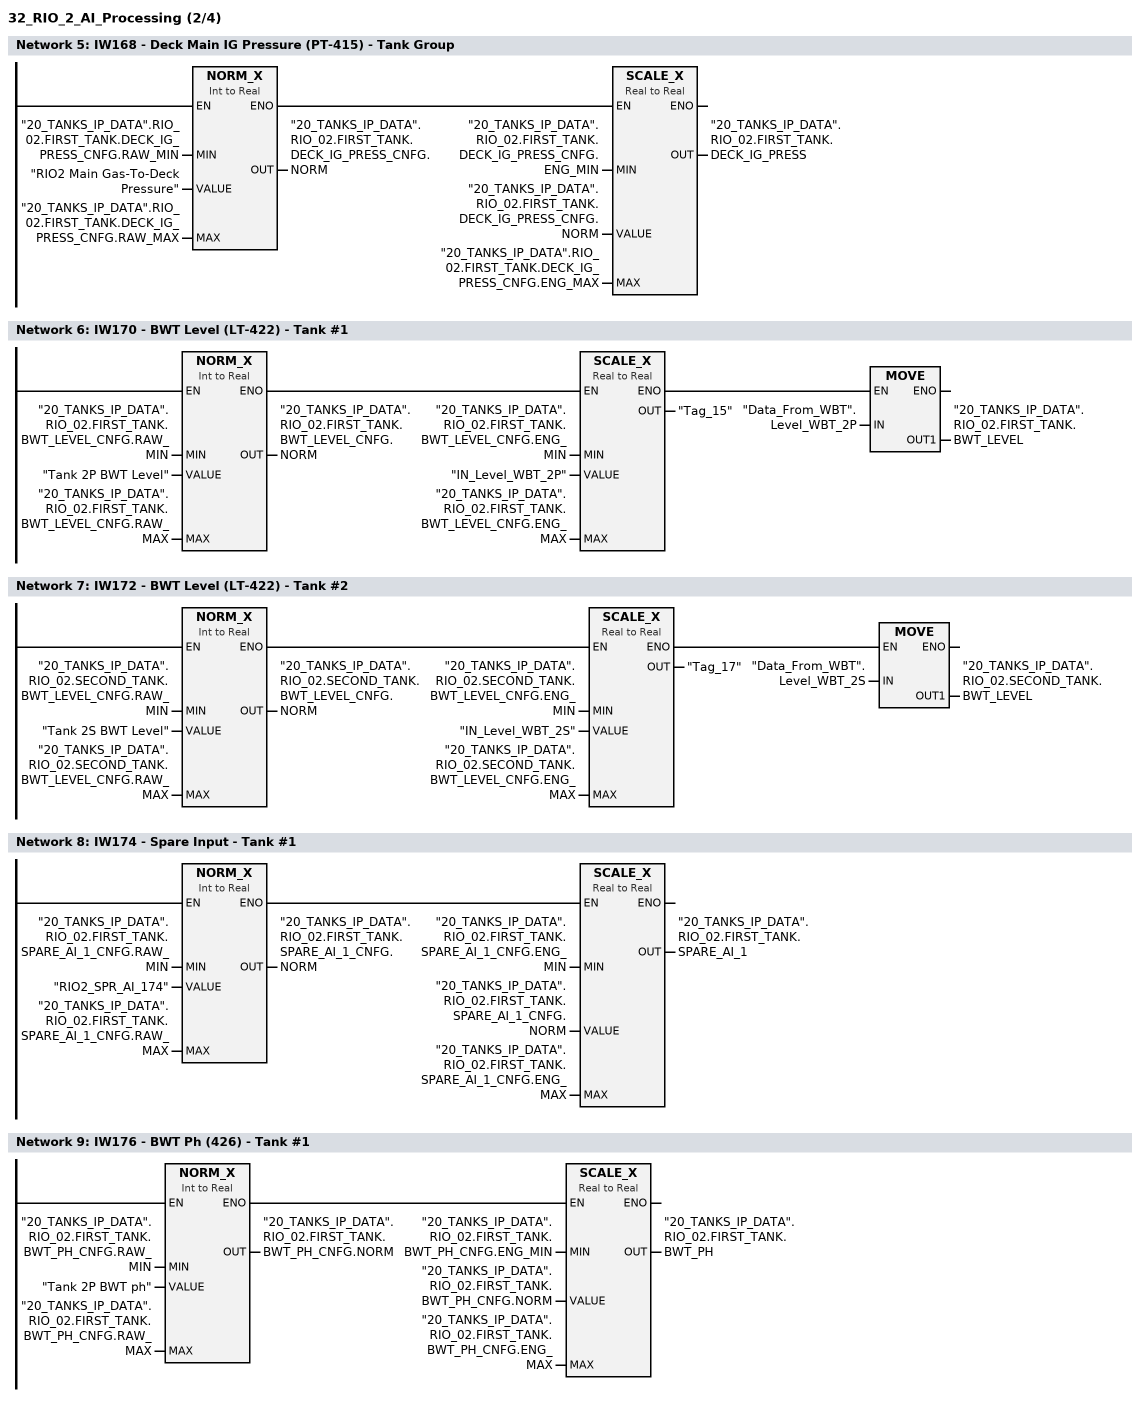
   RUNG wire#powerrail
      { S7_Templates := "[SrcType := Int, DestType := Real]" } Normalize(min := "20_TANKS_IP_DATA".RIO_02.FIRST_TANK.DECK_IG_PRESS_CNFG.RAW_MIN, value := "RIO2 Main Gas-To-Deck Pressure", max := "20_TANKS_IP_DATA".RIO_02.FIRST_TANK.DECK_IG_PRESS_CNFG.RAW_MAX, out => "20_TANKS_IP_DATA".RIO_02.FIRST_TANK.DECK_IG_PRESS_CNFG.NORM)
      { S7_Templates := "[SrcType := Real, DestType := Real]" } Scale(min := "20_TANKS_IP_DATA".RIO_02.FIRST_TANK.DECK_IG_PRESS_CNFG.ENG_MIN, value := "20_TANKS_IP_DATA".RIO_02.FIRST_TANK.DECK_IG_PRESS_CNFG.NORM, max := "20_TANKS_IP_DATA".RIO_02.FIRST_TANK.DECK_IG_PRESS_CNFG.ENG_MAX, out => "20_TANKS_IP_DATA".RIO_02.FIRST_TANK.DECK_IG_PRESS)
   END_RUNG
   // the same network as SCL:
   "20_TANKS_IP_DATA".RIO_02.FIRST_TANK.DECK_IG_PRESS_CNFG.NORM := NORM_X(MIN := "20_TANKS_IP_DATA".RIO_02.FIRST_TANK.DECK_IG_PRESS_CNFG.RAW_MIN, VALUE := "RIO2 Main Gas-To-Deck Pressure", MAX := "20_TANKS_IP_DATA".RIO_02.FIRST_TANK.DECK_IG_PRESS_CNFG.RAW_MAX);
   "20_TANKS_IP_DATA".RIO_02.FIRST_TANK.DECK_IG_PRESS := SCALE_X(MIN := "20_TANKS_IP_DATA".RIO_02.FIRST_TANK.DECK_IG_PRESS_CNFG.ENG_MIN, VALUE := "20_TANKS_IP_DATA".RIO_02.FIRST_TANK.DECK_IG_PRESS_CNFG.NORM, MAX := "20_TANKS_IP_DATA".RIO_02.FIRST_TANK.DECK_IG_PRESS_CNFG.ENG_MAX);
END_REGION

REGION Network 6: IW170 - BWT Level (LT-422) - Tank #1
   RUNG wire#powerrail
      { S7_Templates := "[SrcType := Int, DestType := Real]" } Normalize(min := "20_TANKS_IP_DATA".RIO_02.FIRST_TANK.BWT_LEVEL_CNFG.RAW_MIN, value := "Tank 2P BWT Level", max := "20_TANKS_IP_DATA".RIO_02.FIRST_TANK.BWT_LEVEL_CNFG.RAW_MAX, out => "20_TANKS_IP_DATA".RIO_02.FIRST_TANK.BWT_LEVEL_CNFG.NORM)
      { S7_Templates := "[SrcType := Real, DestType := Real]" } Scale(min := "20_TANKS_IP_DATA".RIO_02.FIRST_TANK.BWT_LEVEL_CNFG.ENG_MIN, value := "IN_Level_WBT_2P", max := "20_TANKS_IP_DATA".RIO_02.FIRST_TANK.BWT_LEVEL_CNFG.ENG_MAX, out => "Tag_15")
      Move(in := "Data_From_WBT".Level_WBT_2P, out1 => "20_TANKS_IP_DATA".RIO_02.FIRST_TANK.BWT_LEVEL)
   END_RUNG
   // the same network as SCL:
   "20_TANKS_IP_DATA".RIO_02.FIRST_TANK.BWT_LEVEL_CNFG.NORM := NORM_X(MIN := "20_TANKS_IP_DATA".RIO_02.FIRST_TANK.BWT_LEVEL_CNFG.RAW_MIN, VALUE := "Tank 2P BWT Level", MAX := "20_TANKS_IP_DATA".RIO_02.FIRST_TANK.BWT_LEVEL_CNFG.RAW_MAX);
   "Tag_15" := SCALE_X(MIN := "20_TANKS_IP_DATA".RIO_02.FIRST_TANK.BWT_LEVEL_CNFG.ENG_MIN, VALUE := "IN_Level_WBT_2P", MAX := "20_TANKS_IP_DATA".RIO_02.FIRST_TANK.BWT_LEVEL_CNFG.ENG_MAX);
   "20_TANKS_IP_DATA".RIO_02.FIRST_TANK.BWT_LEVEL := "Data_From_WBT".Level_WBT_2P;
END_REGION

REGION Network 7: IW172 - BWT Level (LT-422) - Tank #2
   RUNG wire#powerrail
      { S7_Templates := "[SrcType := Int, DestType := Real]" } Normalize(min := "20_TANKS_IP_DATA".RIO_02.SECOND_TANK.BWT_LEVEL_CNFG.RAW_MIN, value := "Tank 2S BWT Level", max := "20_TANKS_IP_DATA".RIO_02.SECOND_TANK.BWT_LEVEL_CNFG.RAW_MAX, out => "20_TANKS_IP_DATA".RIO_02.SECOND_TANK.BWT_LEVEL_CNFG.NORM)
      { S7_Templates := "[SrcType := Real, DestType := Real]" } Scale(min := "20_TANKS_IP_DATA".RIO_02.SECOND_TANK.BWT_LEVEL_CNFG.ENG_MIN, value := "IN_Level_WBT_2S", max := "20_TANKS_IP_DATA".RIO_02.SECOND_TANK.BWT_LEVEL_CNFG.ENG_MAX, out => "Tag_17")
      Move(in := "Data_From_WBT".Level_WBT_2S, out1 => "20_TANKS_IP_DATA".RIO_02.SECOND_TANK.BWT_LEVEL)
   END_RUNG
   // the same network as SCL:
   "20_TANKS_IP_DATA".RIO_02.SECOND_TANK.BWT_LEVEL_CNFG.NORM := NORM_X(MIN := "20_TANKS_IP_DATA".RIO_02.SECOND_TANK.BWT_LEVEL_CNFG.RAW_MIN, VALUE := "Tank 2S BWT Level", MAX := "20_TANKS_IP_DATA".RIO_02.SECOND_TANK.BWT_LEVEL_CNFG.RAW_MAX);
   "Tag_17" := SCALE_X(MIN := "20_TANKS_IP_DATA".RIO_02.SECOND_TANK.BWT_LEVEL_CNFG.ENG_MIN, VALUE := "IN_Level_WBT_2S", MAX := "20_TANKS_IP_DATA".RIO_02.SECOND_TANK.BWT_LEVEL_CNFG.ENG_MAX);
   "20_TANKS_IP_DATA".RIO_02.SECOND_TANK.BWT_LEVEL := "Data_From_WBT".Level_WBT_2S;
END_REGION

REGION Network 8: IW174 - Spare Input - Tank #1
   RUNG wire#powerrail
      { S7_Templates := "[SrcType := Int, DestType := Real]" } Normalize(min := "20_TANKS_IP_DATA".RIO_02.FIRST_TANK.SPARE_AI_1_CNFG.RAW_MIN, value := "RIO2_SPR_AI_174", max := "20_TANKS_IP_DATA".RIO_02.FIRST_TANK.SPARE_AI_1_CNFG.RAW_MAX, out => "20_TANKS_IP_DATA".RIO_02.FIRST_TANK.SPARE_AI_1_CNFG.NORM)
      { S7_Templates := "[SrcType := Real, DestType := Real]" } Scale(min := "20_TANKS_IP_DATA".RIO_02.FIRST_TANK.SPARE_AI_1_CNFG.ENG_MIN, value := "20_TANKS_IP_DATA".RIO_02.FIRST_TANK.SPARE_AI_1_CNFG.NORM, max := "20_TANKS_IP_DATA".RIO_02.FIRST_TANK.SPARE_AI_1_CNFG.ENG_MAX, out => "20_TANKS_IP_DATA".RIO_02.FIRST_TANK.SPARE_AI_1)
   END_RUNG
   // the same network as SCL:
   "20_TANKS_IP_DATA".RIO_02.FIRST_TANK.SPARE_AI_1_CNFG.NORM := NORM_X(MIN := "20_TANKS_IP_DATA".RIO_02.FIRST_TANK.SPARE_AI_1_CNFG.RAW_MIN, VALUE := "RIO2_SPR_AI_174", MAX := "20_TANKS_IP_DATA".RIO_02.FIRST_TANK.SPARE_AI_1_CNFG.RAW_MAX);
   "20_TANKS_IP_DATA".RIO_02.FIRST_TANK.SPARE_AI_1 := SCALE_X(MIN := "20_TANKS_IP_DATA".RIO_02.FIRST_TANK.SPARE_AI_1_CNFG.ENG_MIN, VALUE := "20_TANKS_IP_DATA".RIO_02.FIRST_TANK.SPARE_AI_1_CNFG.NORM, MAX := "20_TANKS_IP_DATA".RIO_02.FIRST_TANK.SPARE_AI_1_CNFG.ENG_MAX);
END_REGION

REGION Network 9: IW176 - BWT Ph (426) - Tank #1
   RUNG wire#powerrail
      { S7_Templates := "[SrcType := Int, DestType := Real]" } Normalize(min := "20_TANKS_IP_DATA".RIO_02.FIRST_TANK.BWT_PH_CNFG.RAW_MIN, value := "Tank 2P BWT ph", max := "20_TANKS_IP_DATA".RIO_02.FIRST_TANK.BWT_PH_CNFG.RAW_MAX, out => "20_TANKS_IP_DATA".RIO_02.FIRST_TANK.BWT_PH_CNFG.NORM)
      { S7_Templates := "[SrcType := Real, DestType := Real]" } Scale(min := "20_TANKS_IP_DATA".RIO_02.FIRST_TANK.BWT_PH_CNFG.ENG_MIN, value := "20_TANKS_IP_DATA".RIO_02.FIRST_TANK.BWT_PH_CNFG.NORM, max := "20_TANKS_IP_DATA".RIO_02.FIRST_TANK.BWT_PH_CNFG.ENG_MAX, out => "20_TANKS_IP_DATA".RIO_02.FIRST_TANK.BWT_PH)
   END_RUNG
   // the same network as SCL:
   "20_TANKS_IP_DATA".RIO_02.FIRST_TANK.BWT_PH_CNFG.NORM := NORM_X(MIN := "20_TANKS_IP_DATA".RIO_02.FIRST_TANK.BWT_PH_CNFG.RAW_MIN, VALUE := "Tank 2P BWT ph", MAX := "20_TANKS_IP_DATA".RIO_02.FIRST_TANK.BWT_PH_CNFG.RAW_MAX);
   "20_TANKS_IP_DATA".RIO_02.FIRST_TANK.BWT_PH := SCALE_X(MIN := "20_TANKS_IP_DATA".RIO_02.FIRST_TANK.BWT_PH_CNFG.ENG_MIN, VALUE := "20_TANKS_IP_DATA".RIO_02.FIRST_TANK.BWT_PH_CNFG.NORM, MAX := "20_TANKS_IP_DATA".RIO_02.FIRST_TANK.BWT_PH_CNFG.ENG_MAX);
END_REGION

REGION Network 10: IW178 - BWT Temperature (426) - Tank #1
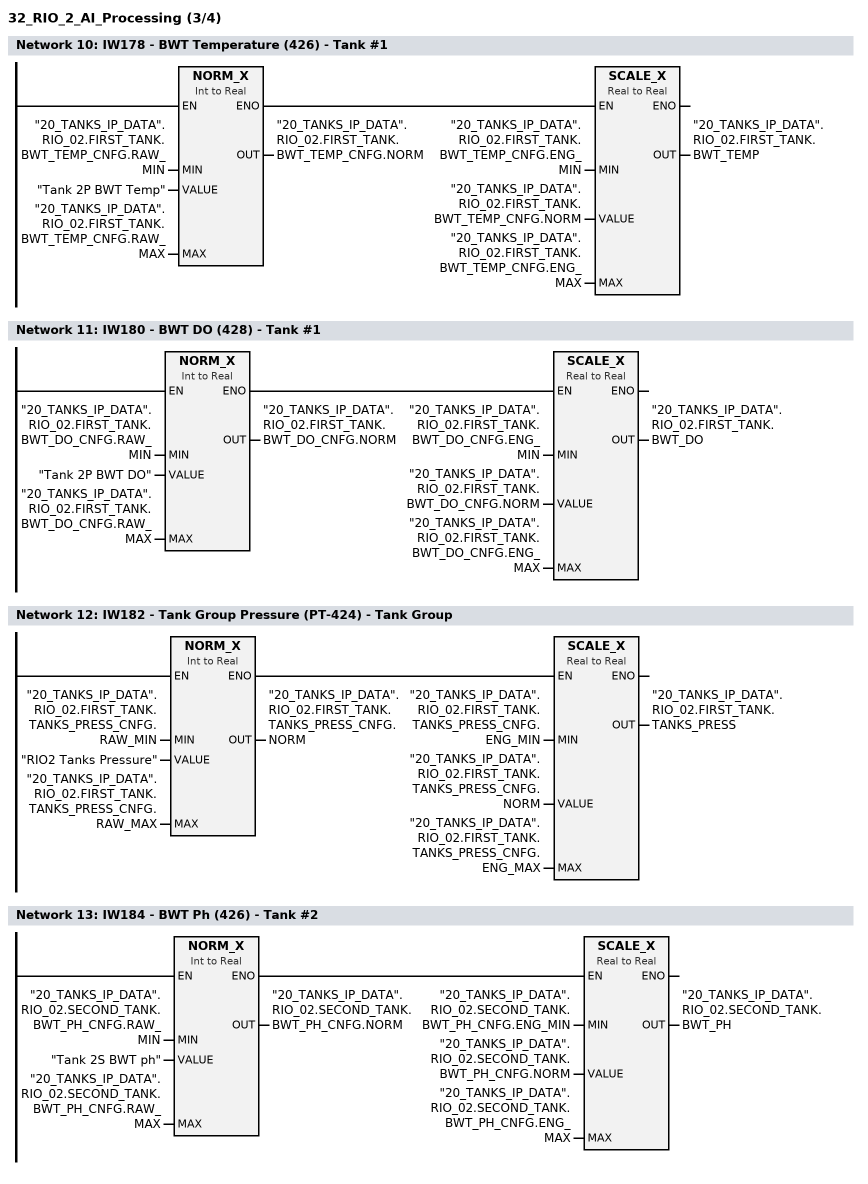
   RUNG wire#powerrail
      { S7_Templates := "[SrcType := Int, DestType := Real]" } Normalize(min := "20_TANKS_IP_DATA".RIO_02.FIRST_TANK.BWT_TEMP_CNFG.RAW_MIN, value := "Tank 2P BWT Temp", max := "20_TANKS_IP_DATA".RIO_02.FIRST_TANK.BWT_TEMP_CNFG.RAW_MAX, out => "20_TANKS_IP_DATA".RIO_02.FIRST_TANK.BWT_TEMP_CNFG.NORM)
      { S7_Templates := "[SrcType := Real, DestType := Real]" } Scale(min := "20_TANKS_IP_DATA".RIO_02.FIRST_TANK.BWT_TEMP_CNFG.ENG_MIN, value := "20_TANKS_IP_DATA".RIO_02.FIRST_TANK.BWT_TEMP_CNFG.NORM, max := "20_TANKS_IP_DATA".RIO_02.FIRST_TANK.BWT_TEMP_CNFG.ENG_MAX, out => "20_TANKS_IP_DATA".RIO_02.FIRST_TANK.BWT_TEMP)
   END_RUNG
   // the same network as SCL:
   "20_TANKS_IP_DATA".RIO_02.FIRST_TANK.BWT_TEMP_CNFG.NORM := NORM_X(MIN := "20_TANKS_IP_DATA".RIO_02.FIRST_TANK.BWT_TEMP_CNFG.RAW_MIN, VALUE := "Tank 2P BWT Temp", MAX := "20_TANKS_IP_DATA".RIO_02.FIRST_TANK.BWT_TEMP_CNFG.RAW_MAX);
   "20_TANKS_IP_DATA".RIO_02.FIRST_TANK.BWT_TEMP := SCALE_X(MIN := "20_TANKS_IP_DATA".RIO_02.FIRST_TANK.BWT_TEMP_CNFG.ENG_MIN, VALUE := "20_TANKS_IP_DATA".RIO_02.FIRST_TANK.BWT_TEMP_CNFG.NORM, MAX := "20_TANKS_IP_DATA".RIO_02.FIRST_TANK.BWT_TEMP_CNFG.ENG_MAX);
END_REGION

REGION Network 11: IW180 - BWT DO (428) - Tank #1
   RUNG wire#powerrail
      { S7_Templates := "[SrcType := Int, DestType := Real]" } Normalize(min := "20_TANKS_IP_DATA".RIO_02.FIRST_TANK.BWT_DO_CNFG.RAW_MIN, value := "Tank 2P BWT DO", max := "20_TANKS_IP_DATA".RIO_02.FIRST_TANK.BWT_DO_CNFG.RAW_MAX, out => "20_TANKS_IP_DATA".RIO_02.FIRST_TANK.BWT_DO_CNFG.NORM)
      { S7_Templates := "[SrcType := Real, DestType := Real]" } Scale(min := "20_TANKS_IP_DATA".RIO_02.FIRST_TANK.BWT_DO_CNFG.ENG_MIN, value := "20_TANKS_IP_DATA".RIO_02.FIRST_TANK.BWT_DO_CNFG.NORM, max := "20_TANKS_IP_DATA".RIO_02.FIRST_TANK.BWT_DO_CNFG.ENG_MAX, out => "20_TANKS_IP_DATA".RIO_02.FIRST_TANK.BWT_DO)
   END_RUNG
   // the same network as SCL:
   "20_TANKS_IP_DATA".RIO_02.FIRST_TANK.BWT_DO_CNFG.NORM := NORM_X(MIN := "20_TANKS_IP_DATA".RIO_02.FIRST_TANK.BWT_DO_CNFG.RAW_MIN, VALUE := "Tank 2P BWT DO", MAX := "20_TANKS_IP_DATA".RIO_02.FIRST_TANK.BWT_DO_CNFG.RAW_MAX);
   "20_TANKS_IP_DATA".RIO_02.FIRST_TANK.BWT_DO := SCALE_X(MIN := "20_TANKS_IP_DATA".RIO_02.FIRST_TANK.BWT_DO_CNFG.ENG_MIN, VALUE := "20_TANKS_IP_DATA".RIO_02.FIRST_TANK.BWT_DO_CNFG.NORM, MAX := "20_TANKS_IP_DATA".RIO_02.FIRST_TANK.BWT_DO_CNFG.ENG_MAX);
END_REGION

REGION Network 12: IW182 - Tank Group Pressure (PT-424) - Tank Group
   RUNG wire#powerrail
      { S7_Templates := "[SrcType := Int, DestType := Real]" } Normalize(min := "20_TANKS_IP_DATA".RIO_02.FIRST_TANK.TANKS_PRESS_CNFG.RAW_MIN, value := "RIO2 Tanks Pressure", max := "20_TANKS_IP_DATA".RIO_02.FIRST_TANK.TANKS_PRESS_CNFG.RAW_MAX, out => "20_TANKS_IP_DATA".RIO_02.FIRST_TANK.TANKS_PRESS_CNFG.NORM)
      { S7_Templates := "[SrcType := Real, DestType := Real]" } Scale(min := "20_TANKS_IP_DATA".RIO_02.FIRST_TANK.TANKS_PRESS_CNFG.ENG_MIN, value := "20_TANKS_IP_DATA".RIO_02.FIRST_TANK.TANKS_PRESS_CNFG.NORM, max := "20_TANKS_IP_DATA".RIO_02.FIRST_TANK.TANKS_PRESS_CNFG.ENG_MAX, out => "20_TANKS_IP_DATA".RIO_02.FIRST_TANK.TANKS_PRESS)
   END_RUNG
   // the same network as SCL:
   "20_TANKS_IP_DATA".RIO_02.FIRST_TANK.TANKS_PRESS_CNFG.NORM := NORM_X(MIN := "20_TANKS_IP_DATA".RIO_02.FIRST_TANK.TANKS_PRESS_CNFG.RAW_MIN, VALUE := "RIO2 Tanks Pressure", MAX := "20_TANKS_IP_DATA".RIO_02.FIRST_TANK.TANKS_PRESS_CNFG.RAW_MAX);
   "20_TANKS_IP_DATA".RIO_02.FIRST_TANK.TANKS_PRESS := SCALE_X(MIN := "20_TANKS_IP_DATA".RIO_02.FIRST_TANK.TANKS_PRESS_CNFG.ENG_MIN, VALUE := "20_TANKS_IP_DATA".RIO_02.FIRST_TANK.TANKS_PRESS_CNFG.NORM, MAX := "20_TANKS_IP_DATA".RIO_02.FIRST_TANK.TANKS_PRESS_CNFG.ENG_MAX);
END_REGION

REGION Network 13: IW184 - BWT Ph (426) - Tank #2
   RUNG wire#powerrail
      { S7_Templates := "[SrcType := Int, DestType := Real]" } Normalize(min := "20_TANKS_IP_DATA".RIO_02.SECOND_TANK.BWT_PH_CNFG.RAW_MIN, value := "Tank 2S BWT ph", max := "20_TANKS_IP_DATA".RIO_02.SECOND_TANK.BWT_PH_CNFG.RAW_MAX, out => "20_TANKS_IP_DATA".RIO_02.SECOND_TANK.BWT_PH_CNFG.NORM)
      { S7_Templates := "[SrcType := Real, DestType := Real]" } Scale(min := "20_TANKS_IP_DATA".RIO_02.SECOND_TANK.BWT_PH_CNFG.ENG_MIN, value := "20_TANKS_IP_DATA".RIO_02.SECOND_TANK.BWT_PH_CNFG.NORM, max := "20_TANKS_IP_DATA".RIO_02.SECOND_TANK.BWT_PH_CNFG.ENG_MAX, out => "20_TANKS_IP_DATA".RIO_02.SECOND_TANK.BWT_PH)
   END_RUNG
   // the same network as SCL:
   "20_TANKS_IP_DATA".RIO_02.SECOND_TANK.BWT_PH_CNFG.NORM := NORM_X(MIN := "20_TANKS_IP_DATA".RIO_02.SECOND_TANK.BWT_PH_CNFG.RAW_MIN, VALUE := "Tank 2S BWT ph", MAX := "20_TANKS_IP_DATA".RIO_02.SECOND_TANK.BWT_PH_CNFG.RAW_MAX);
   "20_TANKS_IP_DATA".RIO_02.SECOND_TANK.BWT_PH := SCALE_X(MIN := "20_TANKS_IP_DATA".RIO_02.SECOND_TANK.BWT_PH_CNFG.ENG_MIN, VALUE := "20_TANKS_IP_DATA".RIO_02.SECOND_TANK.BWT_PH_CNFG.NORM, MAX := "20_TANKS_IP_DATA".RIO_02.SECOND_TANK.BWT_PH_CNFG.ENG_MAX);
END_REGION

REGION Network 14: IW186 - BWT Temperature (426) - Tank #2
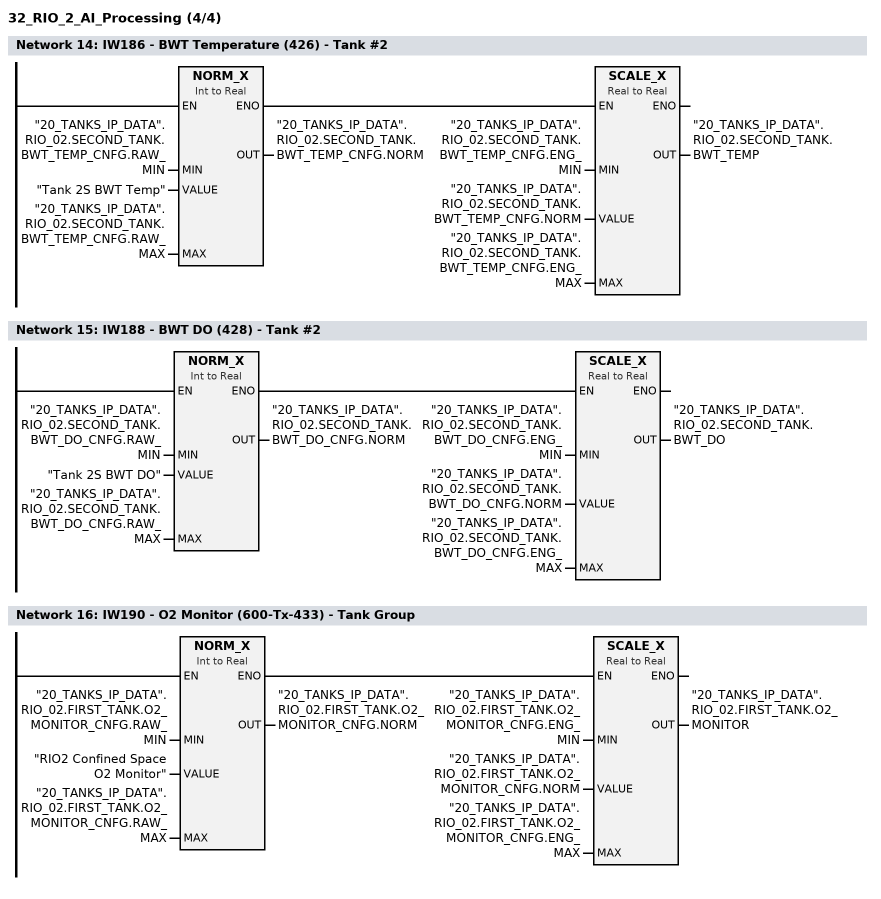
   RUNG wire#powerrail
      { S7_Templates := "[SrcType := Int, DestType := Real]" } Normalize(min := "20_TANKS_IP_DATA".RIO_02.SECOND_TANK.BWT_TEMP_CNFG.RAW_MIN, value := "Tank 2S BWT Temp", max := "20_TANKS_IP_DATA".RIO_02.SECOND_TANK.BWT_TEMP_CNFG.RAW_MAX, out => "20_TANKS_IP_DATA".RIO_02.SECOND_TANK.BWT_TEMP_CNFG.NORM)
      { S7_Templates := "[SrcType := Real, DestType := Real]" } Scale(min := "20_TANKS_IP_DATA".RIO_02.SECOND_TANK.BWT_TEMP_CNFG.ENG_MIN, value := "20_TANKS_IP_DATA".RIO_02.SECOND_TANK.BWT_TEMP_CNFG.NORM, max := "20_TANKS_IP_DATA".RIO_02.SECOND_TANK.BWT_TEMP_CNFG.ENG_MAX, out => "20_TANKS_IP_DATA".RIO_02.SECOND_TANK.BWT_TEMP)
   END_RUNG
   // the same network as SCL:
   "20_TANKS_IP_DATA".RIO_02.SECOND_TANK.BWT_TEMP_CNFG.NORM := NORM_X(MIN := "20_TANKS_IP_DATA".RIO_02.SECOND_TANK.BWT_TEMP_CNFG.RAW_MIN, VALUE := "Tank 2S BWT Temp", MAX := "20_TANKS_IP_DATA".RIO_02.SECOND_TANK.BWT_TEMP_CNFG.RAW_MAX);
   "20_TANKS_IP_DATA".RIO_02.SECOND_TANK.BWT_TEMP := SCALE_X(MIN := "20_TANKS_IP_DATA".RIO_02.SECOND_TANK.BWT_TEMP_CNFG.ENG_MIN, VALUE := "20_TANKS_IP_DATA".RIO_02.SECOND_TANK.BWT_TEMP_CNFG.NORM, MAX := "20_TANKS_IP_DATA".RIO_02.SECOND_TANK.BWT_TEMP_CNFG.ENG_MAX);
END_REGION

REGION Network 15: IW188 - BWT DO (428) - Tank #2
   RUNG wire#powerrail
      { S7_Templates := "[SrcType := Int, DestType := Real]" } Normalize(min := "20_TANKS_IP_DATA".RIO_02.SECOND_TANK.BWT_DO_CNFG.RAW_MIN, value := "Tank 2S BWT DO", max := "20_TANKS_IP_DATA".RIO_02.SECOND_TANK.BWT_DO_CNFG.RAW_MAX, out => "20_TANKS_IP_DATA".RIO_02.SECOND_TANK.BWT_DO_CNFG.NORM)
      { S7_Templates := "[SrcType := Real, DestType := Real]" } Scale(min := "20_TANKS_IP_DATA".RIO_02.SECOND_TANK.BWT_DO_CNFG.ENG_MIN, value := "20_TANKS_IP_DATA".RIO_02.SECOND_TANK.BWT_DO_CNFG.NORM, max := "20_TANKS_IP_DATA".RIO_02.SECOND_TANK.BWT_DO_CNFG.ENG_MAX, out => "20_TANKS_IP_DATA".RIO_02.SECOND_TANK.BWT_DO)
   END_RUNG
   // the same network as SCL:
   "20_TANKS_IP_DATA".RIO_02.SECOND_TANK.BWT_DO_CNFG.NORM := NORM_X(MIN := "20_TANKS_IP_DATA".RIO_02.SECOND_TANK.BWT_DO_CNFG.RAW_MIN, VALUE := "Tank 2S BWT DO", MAX := "20_TANKS_IP_DATA".RIO_02.SECOND_TANK.BWT_DO_CNFG.RAW_MAX);
   "20_TANKS_IP_DATA".RIO_02.SECOND_TANK.BWT_DO := SCALE_X(MIN := "20_TANKS_IP_DATA".RIO_02.SECOND_TANK.BWT_DO_CNFG.ENG_MIN, VALUE := "20_TANKS_IP_DATA".RIO_02.SECOND_TANK.BWT_DO_CNFG.NORM, MAX := "20_TANKS_IP_DATA".RIO_02.SECOND_TANK.BWT_DO_CNFG.ENG_MAX);
END_REGION

REGION Network 16: IW190 - O2 Monitor (600-Tx-433) - Tank Group
   RUNG wire#powerrail
      { S7_Templates := "[SrcType := Int, DestType := Real]" } Normalize(min := "20_TANKS_IP_DATA".RIO_02.FIRST_TANK.O2_MONITOR_CNFG.RAW_MIN, value := "RIO2 Confined Space O2 Monitor", max := "20_TANKS_IP_DATA".RIO_02.FIRST_TANK.O2_MONITOR_CNFG.RAW_MAX, out => "20_TANKS_IP_DATA".RIO_02.FIRST_TANK.O2_MONITOR_CNFG.NORM)
      { S7_Templates := "[SrcType := Real, DestType := Real]" } Scale(min := "20_TANKS_IP_DATA".RIO_02.FIRST_TANK.O2_MONITOR_CNFG.ENG_MIN, value := "20_TANKS_IP_DATA".RIO_02.FIRST_TANK.O2_MONITOR_CNFG.NORM, max := "20_TANKS_IP_DATA".RIO_02.FIRST_TANK.O2_MONITOR_CNFG.ENG_MAX, out => "20_TANKS_IP_DATA".RIO_02.FIRST_TANK.O2_MONITOR)
   END_RUNG
   // the same network as SCL:
   "20_TANKS_IP_DATA".RIO_02.FIRST_TANK.O2_MONITOR_CNFG.NORM := NORM_X(MIN := "20_TANKS_IP_DATA".RIO_02.FIRST_TANK.O2_MONITOR_CNFG.RAW_MIN, VALUE := "RIO2 Confined Space O2 Monitor", MAX := "20_TANKS_IP_DATA".RIO_02.FIRST_TANK.O2_MONITOR_CNFG.RAW_MAX);
   "20_TANKS_IP_DATA".RIO_02.FIRST_TANK.O2_MONITOR := SCALE_X(MIN := "20_TANKS_IP_DATA".RIO_02.FIRST_TANK.O2_MONITOR_CNFG.ENG_MIN, VALUE := "20_TANKS_IP_DATA".RIO_02.FIRST_TANK.O2_MONITOR_CNFG.NORM, MAX := "20_TANKS_IP_DATA".RIO_02.FIRST_TANK.O2_MONITOR_CNFG.ENG_MAX);
END_REGION
END_FUNCTION

FUNCTION "33_RIO_3_AI_Processing" : Void   // FC33, LAD
TITLE = Analogue Input Processing (Tank 1 = 3P, Tank 2 = 3S)
{ S7_Optimized_Access := 'TRUE' }
AUTHOR : JRS
VERSION : 0.1
// To process raw inputs prior to code use
BEGIN

REGION Network 1: IW200 - USD Flow (FIT-418) - Tank #1
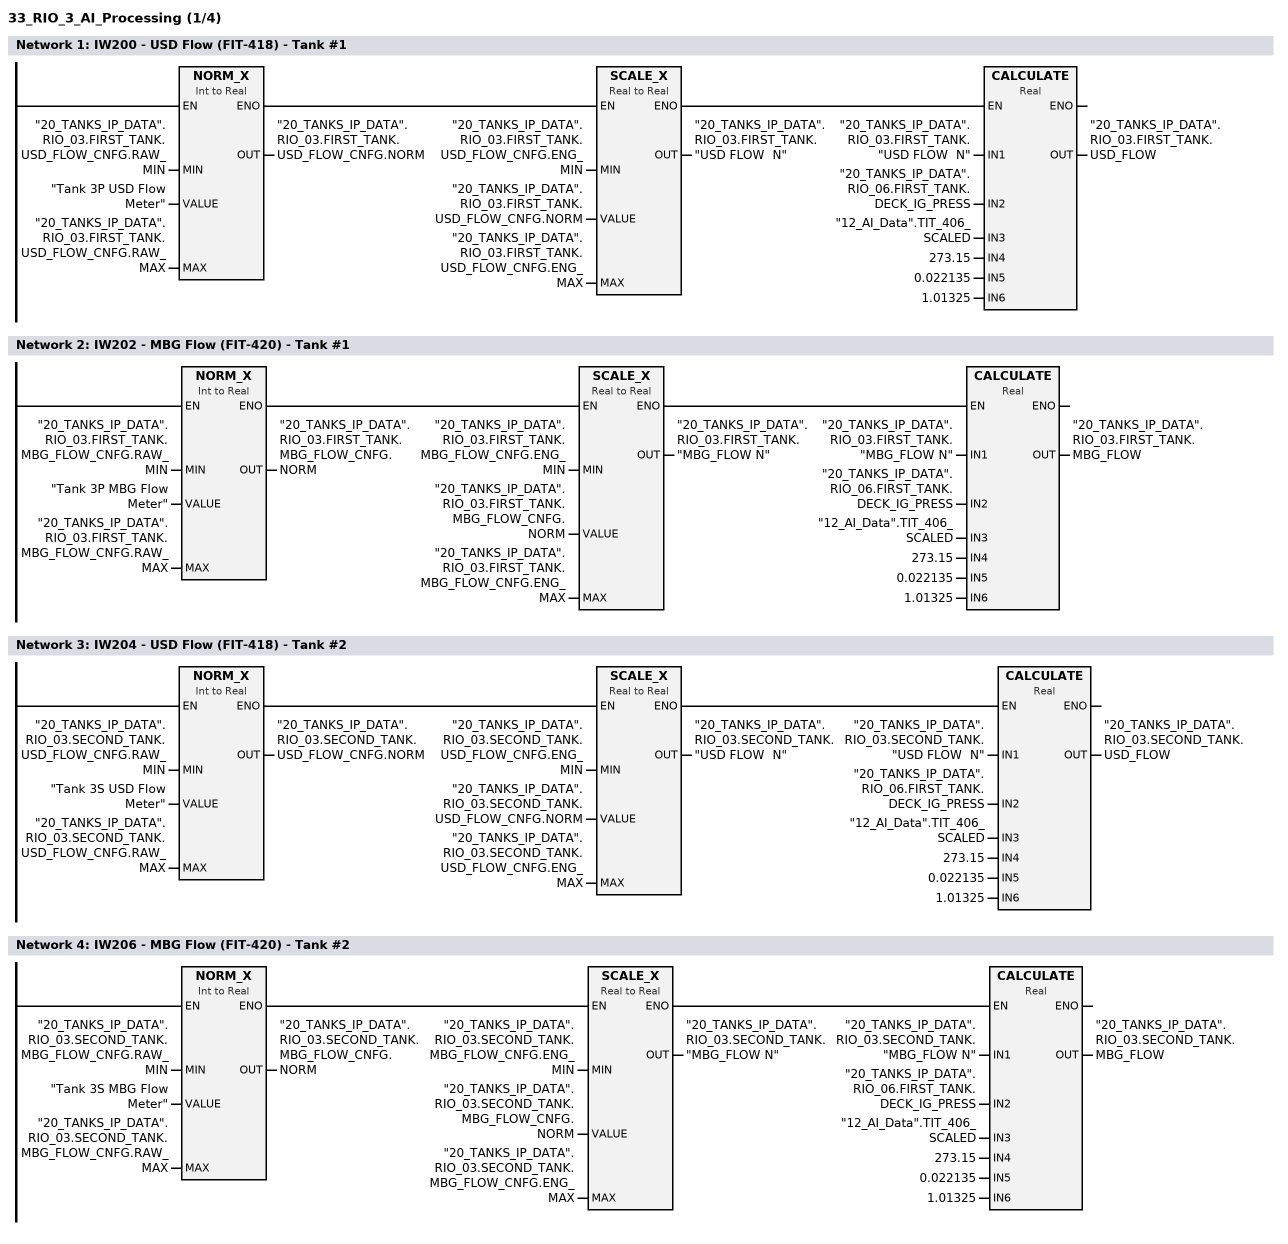
   RUNG wire#powerrail
      { S7_Templates := "[SrcType := Int, DestType := Real]" } Normalize(min := "20_TANKS_IP_DATA".RIO_03.FIRST_TANK.USD_FLOW_CNFG.RAW_MIN, value := "Tank 3P USD Flow Meter", max := "20_TANKS_IP_DATA".RIO_03.FIRST_TANK.USD_FLOW_CNFG.RAW_MAX, out => "20_TANKS_IP_DATA".RIO_03.FIRST_TANK.USD_FLOW_CNFG.NORM)
      { S7_Templates := "[SrcType := Real, DestType := Real]" } Scale(min := "20_TANKS_IP_DATA".RIO_03.FIRST_TANK.USD_FLOW_CNFG.ENG_MIN, value := "20_TANKS_IP_DATA".RIO_03.FIRST_TANK.USD_FLOW_CNFG.NORM, max := "20_TANKS_IP_DATA".RIO_03.FIRST_TANK.USD_FLOW_CNFG.ENG_MAX, out => "20_TANKS_IP_DATA".RIO_03.FIRST_TANK."USD FLOW  N")
      { S7_Templates := "SrcType := Real"; S7_Expression := "IN1*(IN2+IN6)/IN6*IN4/(IN3+IN4)" } Calculate(in1 := "20_TANKS_IP_DATA".RIO_03.FIRST_TANK."USD FLOW  N", in2 := "20_TANKS_IP_DATA".RIO_06.FIRST_TANK.DECK_IG_PRESS, in3 := "12_AI_Data".TIT_406_SCALED, in4 := 273.15, in5 := 0.022135, in6 := 1.01325, out => "20_TANKS_IP_DATA".RIO_03.FIRST_TANK.USD_FLOW)
   END_RUNG
   // the same network as SCL:
   "20_TANKS_IP_DATA".RIO_03.FIRST_TANK.USD_FLOW_CNFG.NORM := NORM_X(MIN := "20_TANKS_IP_DATA".RIO_03.FIRST_TANK.USD_FLOW_CNFG.RAW_MIN, VALUE := "Tank 3P USD Flow Meter", MAX := "20_TANKS_IP_DATA".RIO_03.FIRST_TANK.USD_FLOW_CNFG.RAW_MAX);
   "20_TANKS_IP_DATA".RIO_03.FIRST_TANK."USD FLOW  N" := SCALE_X(MIN := "20_TANKS_IP_DATA".RIO_03.FIRST_TANK.USD_FLOW_CNFG.ENG_MIN, VALUE := "20_TANKS_IP_DATA".RIO_03.FIRST_TANK.USD_FLOW_CNFG.NORM, MAX := "20_TANKS_IP_DATA".RIO_03.FIRST_TANK.USD_FLOW_CNFG.ENG_MAX);
   "20_TANKS_IP_DATA".RIO_03.FIRST_TANK.USD_FLOW := "20_TANKS_IP_DATA".RIO_03.FIRST_TANK."USD FLOW  N"*("20_TANKS_IP_DATA".RIO_06.FIRST_TANK.DECK_IG_PRESS+1.01325)/1.01325*273.15/("12_AI_Data".TIT_406_SCALED+273.15);
END_REGION

REGION Network 2: IW202 - MBG Flow (FIT-420) - Tank #1
   RUNG wire#powerrail
      { S7_Templates := "[SrcType := Int, DestType := Real]" } Normalize(min := "20_TANKS_IP_DATA".RIO_03.FIRST_TANK.MBG_FLOW_CNFG.RAW_MIN, value := "Tank 3P MBG Flow Meter", max := "20_TANKS_IP_DATA".RIO_03.FIRST_TANK.MBG_FLOW_CNFG.RAW_MAX, out => "20_TANKS_IP_DATA".RIO_03.FIRST_TANK.MBG_FLOW_CNFG.NORM)
      { S7_Templates := "[SrcType := Real, DestType := Real]" } Scale(min := "20_TANKS_IP_DATA".RIO_03.FIRST_TANK.MBG_FLOW_CNFG.ENG_MIN, value := "20_TANKS_IP_DATA".RIO_03.FIRST_TANK.MBG_FLOW_CNFG.NORM, max := "20_TANKS_IP_DATA".RIO_03.FIRST_TANK.MBG_FLOW_CNFG.ENG_MAX, out => "20_TANKS_IP_DATA".RIO_03.FIRST_TANK."MBG_FLOW N")
      { S7_Templates := "SrcType := Real"; S7_Expression := "IN1*(IN2+IN6)/IN6*IN4/(IN3+IN4)" } Calculate(in1 := "20_TANKS_IP_DATA".RIO_03.FIRST_TANK."MBG_FLOW N", in2 := "20_TANKS_IP_DATA".RIO_06.FIRST_TANK.DECK_IG_PRESS, in3 := "12_AI_Data".TIT_406_SCALED, in4 := 273.15, in5 := 0.022135, in6 := 1.01325, out => "20_TANKS_IP_DATA".RIO_03.FIRST_TANK.MBG_FLOW)
   END_RUNG
   // the same network as SCL:
   "20_TANKS_IP_DATA".RIO_03.FIRST_TANK.MBG_FLOW_CNFG.NORM := NORM_X(MIN := "20_TANKS_IP_DATA".RIO_03.FIRST_TANK.MBG_FLOW_CNFG.RAW_MIN, VALUE := "Tank 3P MBG Flow Meter", MAX := "20_TANKS_IP_DATA".RIO_03.FIRST_TANK.MBG_FLOW_CNFG.RAW_MAX);
   "20_TANKS_IP_DATA".RIO_03.FIRST_TANK."MBG_FLOW N" := SCALE_X(MIN := "20_TANKS_IP_DATA".RIO_03.FIRST_TANK.MBG_FLOW_CNFG.ENG_MIN, VALUE := "20_TANKS_IP_DATA".RIO_03.FIRST_TANK.MBG_FLOW_CNFG.NORM, MAX := "20_TANKS_IP_DATA".RIO_03.FIRST_TANK.MBG_FLOW_CNFG.ENG_MAX);
   "20_TANKS_IP_DATA".RIO_03.FIRST_TANK.MBG_FLOW := "20_TANKS_IP_DATA".RIO_03.FIRST_TANK."MBG_FLOW N"*("20_TANKS_IP_DATA".RIO_06.FIRST_TANK.DECK_IG_PRESS+1.01325)/1.01325*273.15/("12_AI_Data".TIT_406_SCALED+273.15);
END_REGION

REGION Network 3: IW204 - USD Flow (FIT-418) - Tank #2
   RUNG wire#powerrail
      { S7_Templates := "[SrcType := Int, DestType := Real]" } Normalize(min := "20_TANKS_IP_DATA".RIO_03.SECOND_TANK.USD_FLOW_CNFG.RAW_MIN, value := "Tank 3S USD Flow Meter", max := "20_TANKS_IP_DATA".RIO_03.SECOND_TANK.USD_FLOW_CNFG.RAW_MAX, out => "20_TANKS_IP_DATA".RIO_03.SECOND_TANK.USD_FLOW_CNFG.NORM)
      { S7_Templates := "[SrcType := Real, DestType := Real]" } Scale(min := "20_TANKS_IP_DATA".RIO_03.SECOND_TANK.USD_FLOW_CNFG.ENG_MIN, value := "20_TANKS_IP_DATA".RIO_03.SECOND_TANK.USD_FLOW_CNFG.NORM, max := "20_TANKS_IP_DATA".RIO_03.SECOND_TANK.USD_FLOW_CNFG.ENG_MAX, out => "20_TANKS_IP_DATA".RIO_03.SECOND_TANK."USD FLOW  N")
      { S7_Templates := "SrcType := Real"; S7_Expression := "IN1*(IN2+IN6)/IN6*IN4/(IN3+IN4)" } Calculate(in1 := "20_TANKS_IP_DATA".RIO_03.SECOND_TANK."USD FLOW  N", in2 := "20_TANKS_IP_DATA".RIO_06.FIRST_TANK.DECK_IG_PRESS, in3 := "12_AI_Data".TIT_406_SCALED, in4 := 273.15, in5 := 0.022135, in6 := 1.01325, out => "20_TANKS_IP_DATA".RIO_03.SECOND_TANK.USD_FLOW)
   END_RUNG
   // the same network as SCL:
   "20_TANKS_IP_DATA".RIO_03.SECOND_TANK.USD_FLOW_CNFG.NORM := NORM_X(MIN := "20_TANKS_IP_DATA".RIO_03.SECOND_TANK.USD_FLOW_CNFG.RAW_MIN, VALUE := "Tank 3S USD Flow Meter", MAX := "20_TANKS_IP_DATA".RIO_03.SECOND_TANK.USD_FLOW_CNFG.RAW_MAX);
   "20_TANKS_IP_DATA".RIO_03.SECOND_TANK."USD FLOW  N" := SCALE_X(MIN := "20_TANKS_IP_DATA".RIO_03.SECOND_TANK.USD_FLOW_CNFG.ENG_MIN, VALUE := "20_TANKS_IP_DATA".RIO_03.SECOND_TANK.USD_FLOW_CNFG.NORM, MAX := "20_TANKS_IP_DATA".RIO_03.SECOND_TANK.USD_FLOW_CNFG.ENG_MAX);
   "20_TANKS_IP_DATA".RIO_03.SECOND_TANK.USD_FLOW := "20_TANKS_IP_DATA".RIO_03.SECOND_TANK."USD FLOW  N"*("20_TANKS_IP_DATA".RIO_06.FIRST_TANK.DECK_IG_PRESS+1.01325)/1.01325*273.15/("12_AI_Data".TIT_406_SCALED+273.15);
END_REGION

REGION Network 4: IW206 - MBG Flow (FIT-420) - Tank #2
   RUNG wire#powerrail
      { S7_Templates := "[SrcType := Int, DestType := Real]" } Normalize(min := "20_TANKS_IP_DATA".RIO_03.SECOND_TANK.MBG_FLOW_CNFG.RAW_MIN, value := "Tank 3S MBG Flow Meter", max := "20_TANKS_IP_DATA".RIO_03.SECOND_TANK.MBG_FLOW_CNFG.RAW_MAX, out => "20_TANKS_IP_DATA".RIO_03.SECOND_TANK.MBG_FLOW_CNFG.NORM)
      { S7_Templates := "[SrcType := Real, DestType := Real]" } Scale(min := "20_TANKS_IP_DATA".RIO_03.SECOND_TANK.MBG_FLOW_CNFG.ENG_MIN, value := "20_TANKS_IP_DATA".RIO_03.SECOND_TANK.MBG_FLOW_CNFG.NORM, max := "20_TANKS_IP_DATA".RIO_03.SECOND_TANK.MBG_FLOW_CNFG.ENG_MAX, out => "20_TANKS_IP_DATA".RIO_03.SECOND_TANK."MBG_FLOW N")
      { S7_Templates := "SrcType := Real"; S7_Expression := "IN1*(IN2+IN6)/IN6*IN4/(IN3+IN4)" } Calculate(in1 := "20_TANKS_IP_DATA".RIO_03.SECOND_TANK."MBG_FLOW N", in2 := "20_TANKS_IP_DATA".RIO_06.FIRST_TANK.DECK_IG_PRESS, in3 := "12_AI_Data".TIT_406_SCALED, in4 := 273.15, in5 := 0.022135, in6 := 1.01325, out => "20_TANKS_IP_DATA".RIO_03.SECOND_TANK.MBG_FLOW)
   END_RUNG
   // the same network as SCL:
   "20_TANKS_IP_DATA".RIO_03.SECOND_TANK.MBG_FLOW_CNFG.NORM := NORM_X(MIN := "20_TANKS_IP_DATA".RIO_03.SECOND_TANK.MBG_FLOW_CNFG.RAW_MIN, VALUE := "Tank 3S MBG Flow Meter", MAX := "20_TANKS_IP_DATA".RIO_03.SECOND_TANK.MBG_FLOW_CNFG.RAW_MAX);
   "20_TANKS_IP_DATA".RIO_03.SECOND_TANK."MBG_FLOW N" := SCALE_X(MIN := "20_TANKS_IP_DATA".RIO_03.SECOND_TANK.MBG_FLOW_CNFG.ENG_MIN, VALUE := "20_TANKS_IP_DATA".RIO_03.SECOND_TANK.MBG_FLOW_CNFG.NORM, MAX := "20_TANKS_IP_DATA".RIO_03.SECOND_TANK.MBG_FLOW_CNFG.ENG_MAX);
   "20_TANKS_IP_DATA".RIO_03.SECOND_TANK.MBG_FLOW := "20_TANKS_IP_DATA".RIO_03.SECOND_TANK."MBG_FLOW N"*("20_TANKS_IP_DATA".RIO_06.FIRST_TANK.DECK_IG_PRESS+1.01325)/1.01325*273.15/("12_AI_Data".TIT_406_SCALED+273.15);
END_REGION

REGION Network 5: IW208 - Deck Main IG Pressure (PT-415) - Tank Group
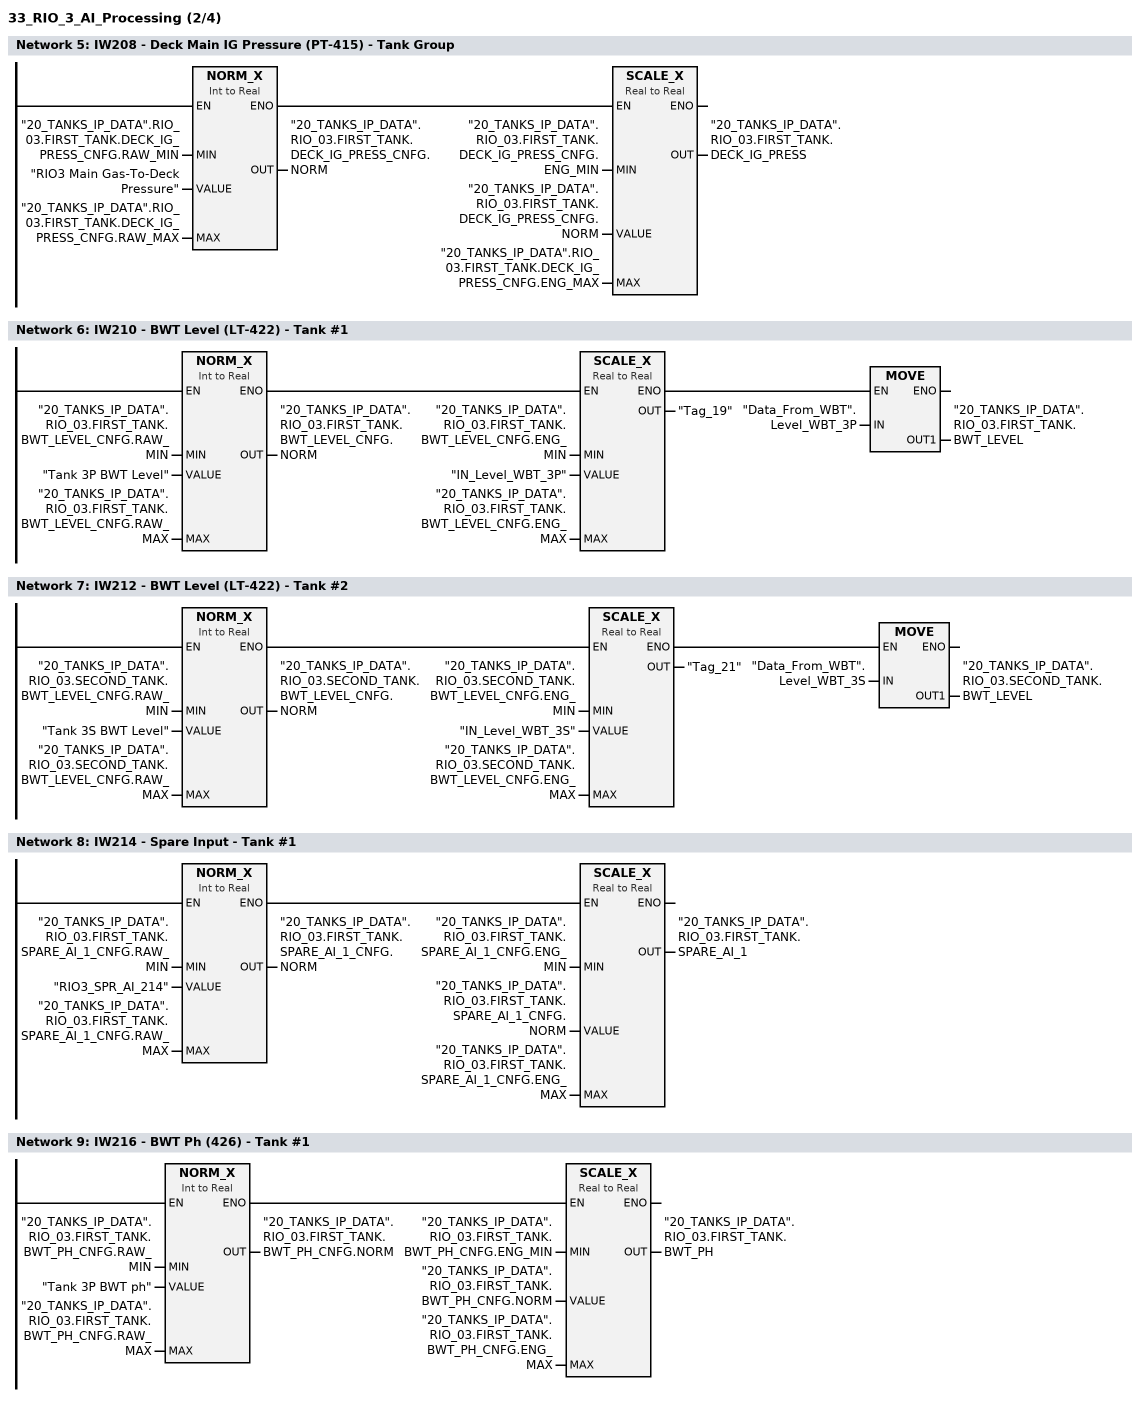
   RUNG wire#powerrail
      { S7_Templates := "[SrcType := Int, DestType := Real]" } Normalize(min := "20_TANKS_IP_DATA".RIO_03.FIRST_TANK.DECK_IG_PRESS_CNFG.RAW_MIN, value := "RIO3 Main Gas-To-Deck Pressure", max := "20_TANKS_IP_DATA".RIO_03.FIRST_TANK.DECK_IG_PRESS_CNFG.RAW_MAX, out => "20_TANKS_IP_DATA".RIO_03.FIRST_TANK.DECK_IG_PRESS_CNFG.NORM)
      { S7_Templates := "[SrcType := Real, DestType := Real]" } Scale(min := "20_TANKS_IP_DATA".RIO_03.FIRST_TANK.DECK_IG_PRESS_CNFG.ENG_MIN, value := "20_TANKS_IP_DATA".RIO_03.FIRST_TANK.DECK_IG_PRESS_CNFG.NORM, max := "20_TANKS_IP_DATA".RIO_03.FIRST_TANK.DECK_IG_PRESS_CNFG.ENG_MAX, out => "20_TANKS_IP_DATA".RIO_03.FIRST_TANK.DECK_IG_PRESS)
   END_RUNG
   // the same network as SCL:
   "20_TANKS_IP_DATA".RIO_03.FIRST_TANK.DECK_IG_PRESS_CNFG.NORM := NORM_X(MIN := "20_TANKS_IP_DATA".RIO_03.FIRST_TANK.DECK_IG_PRESS_CNFG.RAW_MIN, VALUE := "RIO3 Main Gas-To-Deck Pressure", MAX := "20_TANKS_IP_DATA".RIO_03.FIRST_TANK.DECK_IG_PRESS_CNFG.RAW_MAX);
   "20_TANKS_IP_DATA".RIO_03.FIRST_TANK.DECK_IG_PRESS := SCALE_X(MIN := "20_TANKS_IP_DATA".RIO_03.FIRST_TANK.DECK_IG_PRESS_CNFG.ENG_MIN, VALUE := "20_TANKS_IP_DATA".RIO_03.FIRST_TANK.DECK_IG_PRESS_CNFG.NORM, MAX := "20_TANKS_IP_DATA".RIO_03.FIRST_TANK.DECK_IG_PRESS_CNFG.ENG_MAX);
END_REGION

